REGION Network 3: I75.2 - Tank Vent Valve 1 Feedback Open (CV-441-A)
   // True = OPEN, False = NOT
   RUNG wire#powerrail
      Contact( "APT Tank Vent Valve 1 Feedback - Opened" )
      Coil( "20_TANKS_IP_DATA".RIO_07.FIRST_TANK.TANK_VENT_A_OPEN )
   END_RUNG
   // the same network as SCL:
   "20_TANKS_IP_DATA".RIO_07.FIRST_TANK.TANK_VENT_A_OPEN := "APT Tank Vent Valve 1 Feedback - Opened";
END_REGION

REGION Network 4: I75.3 - Tank Vent Valve 1 Feedback Closed (CV-441-A)
   // True = CLOSED, False = NOT
   RUNG wire#powerrail
      Contact( "APT Tank Vent Valve 1 Feedback - Closed" )
      Coil( "20_TANKS_IP_DATA".RIO_07.FIRST_TANK.TANK_VENT_A_CLSD )
   END_RUNG
   // the same network as SCL:
   "20_TANKS_IP_DATA".RIO_07.FIRST_TANK.TANK_VENT_A_CLSD := "APT Tank Vent Valve 1 Feedback - Closed";
END_REGION

REGION Network 5: I75.4 - Tank Vent Valve 2 Feedback Open (CV-441-B)
   // True = OPEN, False = NOT
   RUNG wire#powerrail
      Contact( "APT Tank Vent Valve 2 Feedback - Opened" )
      Coil( "20_TANKS_IP_DATA".RIO_07.FIRST_TANK.TANK_VENT_B_OPEN )
   END_RUNG
   // the same network as SCL:
   "20_TANKS_IP_DATA".RIO_07.FIRST_TANK.TANK_VENT_B_OPEN := "APT Tank Vent Valve 2 Feedback - Opened";
END_REGION

REGION Network 6: I75.5 - Tank Vent Valve 2 Feedback Closed (CV-441-B)
   // True = CLOSED, False = NOT
   RUNG wire#powerrail
      Contact( "APT Tank Vent Valve 2 Feedback - Closed" )
      Coil( "20_TANKS_IP_DATA".RIO_07.FIRST_TANK.TANK_VENT_B_CLSD )
   END_RUNG
   // the same network as SCL:
   "20_TANKS_IP_DATA".RIO_07.FIRST_TANK.TANK_VENT_B_CLSD := "APT Tank Vent Valve 2 Feedback - Closed";
END_REGION

REGION Network 7: I75.6 - Spare Input Destination Accesed from Warning FC
   // True = N/A, False = N/A
END_REGION

REGION Network 8: I75.7 - Spare Input
   // True = N/A, False = N/A
   RUNG wire#powerrail
      Contact( "RIO7_SPR_DI_175_7" )
      Coil( "20_TANKS_IP_DATA".RIO_07.FIRST_TANK.SPARE_DI_7 )
   END_RUNG
   // the same network as SCL:
   "20_TANKS_IP_DATA".RIO_07.FIRST_TANK.SPARE_DI_7 := "RIO7_SPR_DI_175_7";
END_REGION

REGION Network 9: I78.0 - Tank Level HIHI - (LS-425) - First Tank
   // True = OK, False = HIHI
   RUNG wire#powerrail
      I_Contact( "APT BWT Level High High Switch" )
      Coil( "20_TANKS_IP_DATA".RIO_07.FIRST_TANK.BWT_LEVEL_HIHI )
   END_RUNG
   // the same network as SCL:
   "20_TANKS_IP_DATA".RIO_07.FIRST_TANK.BWT_LEVEL_HIHI := NOT "APT BWT Level High High Switch";
END_REGION

REGION Network 10: I78.1 - Tank Group Pressure HIHI (PS-436)
   // True = OK, False = HIHI
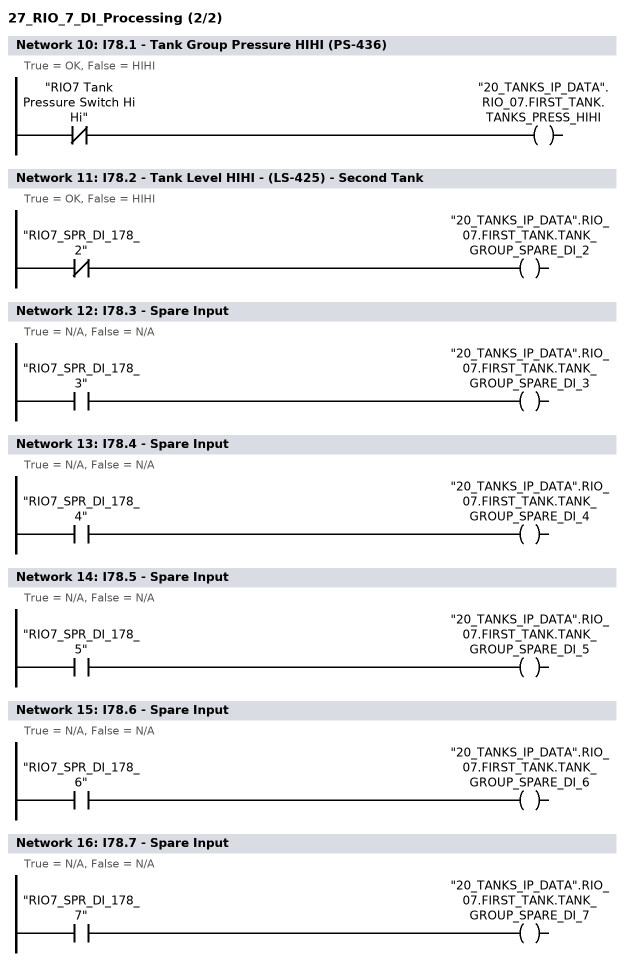
   RUNG wire#powerrail
      I_Contact( "RIO7 Tank Pressure Switch Hi Hi" )
      Coil( "20_TANKS_IP_DATA".RIO_07.FIRST_TANK.TANKS_PRESS_HIHI )
   END_RUNG
   // the same network as SCL:
   "20_TANKS_IP_DATA".RIO_07.FIRST_TANK.TANKS_PRESS_HIHI := NOT "RIO7 Tank Pressure Switch Hi Hi";
END_REGION

REGION Network 11: I78.2 - Tank Level HIHI - (LS-425) - Second Tank
   // True = OK, False = HIHI
   RUNG wire#powerrail
      I_Contact( "RIO7_SPR_DI_178_2" )
      Coil( "20_TANKS_IP_DATA".RIO_07.FIRST_TANK.TANK_GROUP_SPARE_DI_2 )
   END_RUNG
   // the same network as SCL:
   "20_TANKS_IP_DATA".RIO_07.FIRST_TANK.TANK_GROUP_SPARE_DI_2 := NOT "RIO7_SPR_DI_178_2";
END_REGION

REGION Network 12: I78.3 - Spare Input
   // True = N/A, False = N/A
   RUNG wire#powerrail
      Contact( "RIO7_SPR_DI_178_3" )
      Coil( "20_TANKS_IP_DATA".RIO_07.FIRST_TANK.TANK_GROUP_SPARE_DI_3 )
   END_RUNG
   // the same network as SCL:
   "20_TANKS_IP_DATA".RIO_07.FIRST_TANK.TANK_GROUP_SPARE_DI_3 := "RIO7_SPR_DI_178_3";
END_REGION

REGION Network 13: I78.4 - Spare Input
   // True = N/A, False = N/A
   RUNG wire#powerrail
      Contact( "RIO7_SPR_DI_178_4" )
      Coil( "20_TANKS_IP_DATA".RIO_07.FIRST_TANK.TANK_GROUP_SPARE_DI_4 )
   END_RUNG
   // the same network as SCL:
   "20_TANKS_IP_DATA".RIO_07.FIRST_TANK.TANK_GROUP_SPARE_DI_4 := "RIO7_SPR_DI_178_4";
END_REGION

REGION Network 14: I78.5 - Spare Input
   // True = N/A, False = N/A
   RUNG wire#powerrail
      Contact( "RIO7_SPR_DI_178_5" )
      Coil( "20_TANKS_IP_DATA".RIO_07.FIRST_TANK.TANK_GROUP_SPARE_DI_5 )
   END_RUNG
   // the same network as SCL:
   "20_TANKS_IP_DATA".RIO_07.FIRST_TANK.TANK_GROUP_SPARE_DI_5 := "RIO7_SPR_DI_178_5";
END_REGION

REGION Network 15: I78.6 - Spare Input
   // True = N/A, False = N/A
   RUNG wire#powerrail
      Contact( "RIO7_SPR_DI_178_6" )
      Coil( "20_TANKS_IP_DATA".RIO_07.FIRST_TANK.TANK_GROUP_SPARE_DI_6 )
   END_RUNG
   // the same network as SCL:
   "20_TANKS_IP_DATA".RIO_07.FIRST_TANK.TANK_GROUP_SPARE_DI_6 := "RIO7_SPR_DI_178_6";
END_REGION

REGION Network 16: I78.7 - Spare Input
   // True = N/A, False = N/A
   RUNG wire#powerrail
      Contact( "RIO7_SPR_DI_178_7" )
      Coil( "20_TANKS_IP_DATA".RIO_07.FIRST_TANK.TANK_GROUP_SPARE_DI_7 )
   END_RUNG
   // the same network as SCL:
   "20_TANKS_IP_DATA".RIO_07.FIRST_TANK.TANK_GROUP_SPARE_DI_7 := "RIO7_SPR_DI_178_7";
END_REGION
END_FUNCTION

FUNCTION "WBTs" : Void   // FC28, SCL
{ S7_Optimized_Access := 'TRUE' }
VERSION : 0.1
BEGIN
   "Data_From_WBT"."Level_FPT" := (INT_TO_REAL("IN_Level_FPT") / 1000.0) / "Data_From_WBT".Level_Max_FPT * 100.0;
   "Data_From_WBT"."Level_FPT m" := (INT_TO_REAL("IN_Level_FPT") / 1000.0);

   "Data_From_WBT"."Level_WBT_1S" := (INT_TO_REAL("IN_Level_WBT_1S") / 1000.0) /"Data_From_WBT".Level_Max_WBT_1S * 100.0;
   "Data_From_WBT"."Level_WBT_1P" := (INT_TO_REAL("IN_Level_WBT_1P") / 1000.0) / "Data_From_WBT".Level_Max_WBT_1P * 100.0;
   "Data_From_WBT"."Level_WBT_1S m" := (INT_TO_REAL("IN_Level_WBT_1S") / 1000.0);
   "Data_From_WBT"."Level_WBT_1P m" := (INT_TO_REAL("IN_Level_WBT_1P") / 1000.0);

   "Data_From_WBT"."Level_WBT_2S" := (INT_TO_REAL("IN_Level_WBT_2S") / 1000.0) / "Data_From_WBT".Level_Max_WBT_2S * 100.0;
   "Data_From_WBT"."Level_WBT_2P" := (INT_TO_REAL("IN_Level_WBT_2P") / 1000.0) / "Data_From_WBT".Level_Max_WBT_2P * 100.0;
   "Data_From_WBT"."Level_WBT_2S m":= (INT_TO_REAL("IN_Level_WBT_2S") / 1000.0);
   "Data_From_WBT"."Level_WBT_2P m" := (INT_TO_REAL("IN_Level_WBT_2P") / 1000.0);

   "Data_From_WBT"."Level_WBT_3S" := (INT_TO_REAL("IN_Level_WBT_3S") / 1000.0) / "Data_From_WBT".Level_Max_WBT_3S * 100.0;
   "Data_From_WBT"."Level_WBT_3P" := (INT_TO_REAL("IN_Level_WBT_3P") / 1000.0) / "Data_From_WBT".Level_Max_WBT_3P * 100.0;
   "Data_From_WBT"."Level_WBT_3S m" := (INT_TO_REAL("IN_Level_WBT_3S") / 1000.0);
   "Data_From_WBT"."Level_WBT_3P m" := (INT_TO_REAL("IN_Level_WBT_3P") / 1000.0);

   "Data_From_WBT"."Level_WBT_4S" := (INT_TO_REAL("IN_Level_WBT_4S") / 1000.0) / "Data_From_WBT".Level_Max_WBT_4S * 100.0;
   "Data_From_WBT"."Level_WBT_4P" := (INT_TO_REAL("IN_Level_WBT_4P") / 1000.0) / "Data_From_WBT".Level_Max_WBT_4P * 100.0;
   "Data_From_WBT"."Level_WBT_4S m" := (INT_TO_REAL("IN_Level_WBT_4S") / 1000.0);
   "Data_From_WBT"."Level_WBT_4P m" := (INT_TO_REAL("IN_Level_WBT_4P") / 1000.0);

   "Data_From_WBT"."Level_WBT_5S" := (INT_TO_REAL("IN_Level_WBT_5S") / 1000.0) / "Data_From_WBT".Level_Max_WBT_5S * 100.0;
   "Data_From_WBT"."Level_WBT_5P" := (INT_TO_REAL("IN_Level_WBT_5P") / 1000.0) / "Data_From_WBT".Level_Max_WBT_5P * 100.0;
   "Data_From_WBT"."Level_WBT_5S m" := (INT_TO_REAL("IN_Level_WBT_5S") / 1000.0);
   "Data_From_WBT"."Level_WBT_5P m" := (INT_TO_REAL("IN_Level_WBT_5P") / 1000.0);

   "Data_From_WBT"."Level_WBT_6S" := (INT_TO_REAL("IN_Level_WBT_6S") / 1000.0) / "Data_From_WBT".Level_Max_WBT_6S * 100.0;
   "Data_From_WBT"."Level_WBT_6P" := (INT_TO_REAL("IN_Level_WBT_6P") / 1000.0) / "Data_From_WBT".Level_Max_WBT_6P * 100.0;
   "Data_From_WBT"."Level_WBT_6S m" := (INT_TO_REAL("IN_Level_WBT_6S") / 1000.0);
   "Data_From_WBT"."Level_WBT_6P m" := (INT_TO_REAL("IN_Level_WBT_6P") / 1000.0);

   "Data_From_WBT"."Level_APT" := (INT_TO_REAL("IN_Level_APT") / 1000.0) / "Data_From_WBT".Level_Max_APT * 100.0;
   "Data_From_WBT"."Level_APT m" := (INT_TO_REAL("IN_Level_APT") / 1000.0);
END_FUNCTION

FUNCTION "31_RIO_1_AI_Processing" : Void   // FC31, LAD
TITLE = Analogue Input Processing (Tank 1 = FPT, Tank 2 = 1P, Tank 3 = 1S)
{ S7_Optimized_Access := 'TRUE' }
AUTHOR : JRS
VERSION : 0.1
// To process raw inputs prior to code use
BEGIN

REGION Network 1: IW100 - USD Flow (FIT-418) - Tank #1
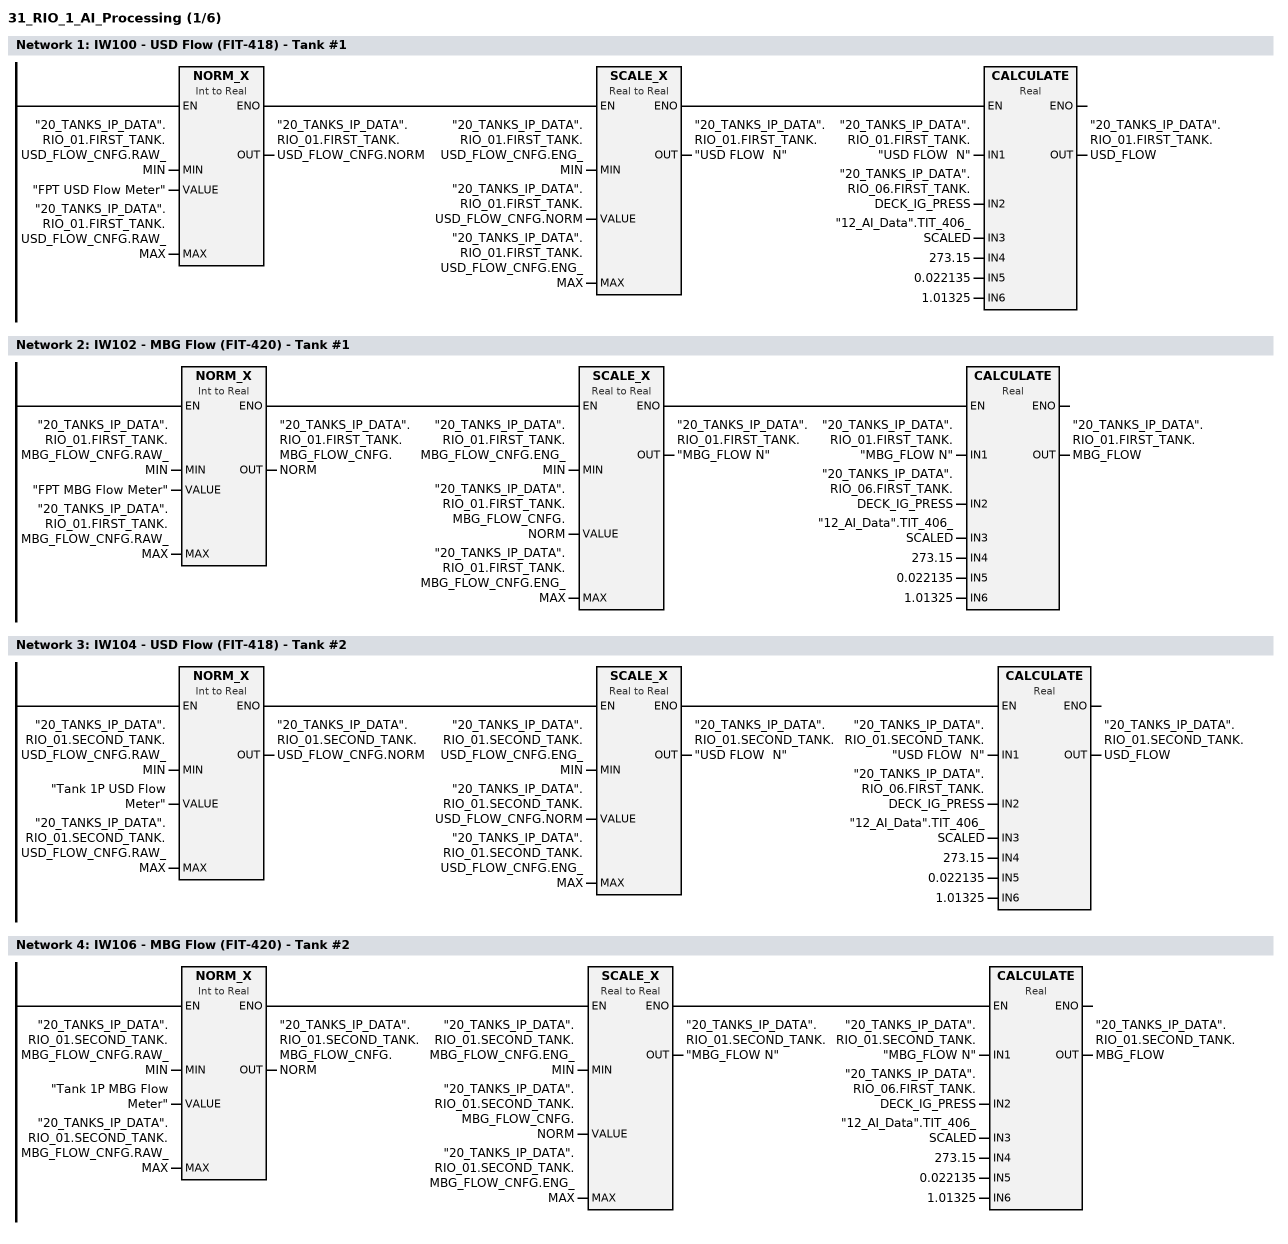
   RUNG wire#powerrail
      { S7_Templates := "[SrcType := Int, DestType := Real]" } Normalize(min := "20_TANKS_IP_DATA".RIO_01.FIRST_TANK.USD_FLOW_CNFG.RAW_MIN, value := "FPT USD Flow Meter", max := "20_TANKS_IP_DATA".RIO_01.FIRST_TANK.USD_FLOW_CNFG.RAW_MAX, out => "20_TANKS_IP_DATA".RIO_01.FIRST_TANK.USD_FLOW_CNFG.NORM)
      { S7_Templates := "[SrcType := Real, DestType := Real]" } Scale(min := "20_TANKS_IP_DATA".RIO_01.FIRST_TANK.USD_FLOW_CNFG.ENG_MIN, value := "20_TANKS_IP_DATA".RIO_01.FIRST_TANK.USD_FLOW_CNFG.NORM, max := "20_TANKS_IP_DATA".RIO_01.FIRST_TANK.USD_FLOW_CNFG.ENG_MAX, out => "20_TANKS_IP_DATA".RIO_01.FIRST_TANK."USD FLOW  N")
      { S7_Templates := "SrcType := Real"; S7_Expression := "IN1*(IN2+IN6)/IN6*IN4/(IN3+IN4)" } Calculate(in1 := "20_TANKS_IP_DATA".RIO_01.FIRST_TANK."USD FLOW  N", in2 := "20_TANKS_IP_DATA".RIO_06.FIRST_TANK.DECK_IG_PRESS, in3 := "12_AI_Data".TIT_406_SCALED, in4 := 273.15, in5 := 0.022135, in6 := 1.01325, out => "20_TANKS_IP_DATA".RIO_01.FIRST_TANK.USD_FLOW)
   END_RUNG
   // the same network as SCL:
   "20_TANKS_IP_DATA".RIO_01.FIRST_TANK.USD_FLOW_CNFG.NORM := NORM_X(MIN := "20_TANKS_IP_DATA".RIO_01.FIRST_TANK.USD_FLOW_CNFG.RAW_MIN, VALUE := "FPT USD Flow Meter", MAX := "20_TANKS_IP_DATA".RIO_01.FIRST_TANK.USD_FLOW_CNFG.RAW_MAX);
   "20_TANKS_IP_DATA".RIO_01.FIRST_TANK."USD FLOW  N" := SCALE_X(MIN := "20_TANKS_IP_DATA".RIO_01.FIRST_TANK.USD_FLOW_CNFG.ENG_MIN, VALUE := "20_TANKS_IP_DATA".RIO_01.FIRST_TANK.USD_FLOW_CNFG.NORM, MAX := "20_TANKS_IP_DATA".RIO_01.FIRST_TANK.USD_FLOW_CNFG.ENG_MAX);
   "20_TANKS_IP_DATA".RIO_01.FIRST_TANK.USD_FLOW := "20_TANKS_IP_DATA".RIO_01.FIRST_TANK."USD FLOW  N"*("20_TANKS_IP_DATA".RIO_06.FIRST_TANK.DECK_IG_PRESS+1.01325)/1.01325*273.15/("12_AI_Data".TIT_406_SCALED+273.15);
END_REGION

REGION Network 2: IW102 - MBG Flow (FIT-420) - Tank #1
   RUNG wire#powerrail
      { S7_Templates := "[SrcType := Int, DestType := Real]" } Normalize(min := "20_TANKS_IP_DATA".RIO_01.FIRST_TANK.MBG_FLOW_CNFG.RAW_MIN, value := "FPT MBG Flow Meter", max := "20_TANKS_IP_DATA".RIO_01.FIRST_TANK.MBG_FLOW_CNFG.RAW_MAX, out => "20_TANKS_IP_DATA".RIO_01.FIRST_TANK.MBG_FLOW_CNFG.NORM)
      { S7_Templates := "[SrcType := Real, DestType := Real]" } Scale(min := "20_TANKS_IP_DATA".RIO_01.FIRST_TANK.MBG_FLOW_CNFG.ENG_MIN, value := "20_TANKS_IP_DATA".RIO_01.FIRST_TANK.MBG_FLOW_CNFG.NORM, max := "20_TANKS_IP_DATA".RIO_01.FIRST_TANK.MBG_FLOW_CNFG.ENG_MAX, out => "20_TANKS_IP_DATA".RIO_01.FIRST_TANK."MBG_FLOW N")
      { S7_Templates := "SrcType := Real"; S7_Expression := "IN1*(IN2+IN6)/IN6*IN4/(IN3+IN4)" } Calculate(in1 := "20_TANKS_IP_DATA".RIO_01.FIRST_TANK."MBG_FLOW N", in2 := "20_TANKS_IP_DATA".RIO_06.FIRST_TANK.DECK_IG_PRESS, in3 := "12_AI_Data".TIT_406_SCALED, in4 := 273.15, in5 := 0.022135, in6 := 1.01325, out => "20_TANKS_IP_DATA".RIO_01.FIRST_TANK.MBG_FLOW)
   END_RUNG
   // the same network as SCL:
   "20_TANKS_IP_DATA".RIO_01.FIRST_TANK.MBG_FLOW_CNFG.NORM := NORM_X(MIN := "20_TANKS_IP_DATA".RIO_01.FIRST_TANK.MBG_FLOW_CNFG.RAW_MIN, VALUE := "FPT MBG Flow Meter", MAX := "20_TANKS_IP_DATA".RIO_01.FIRST_TANK.MBG_FLOW_CNFG.RAW_MAX);
   "20_TANKS_IP_DATA".RIO_01.FIRST_TANK."MBG_FLOW N" := SCALE_X(MIN := "20_TANKS_IP_DATA".RIO_01.FIRST_TANK.MBG_FLOW_CNFG.ENG_MIN, VALUE := "20_TANKS_IP_DATA".RIO_01.FIRST_TANK.MBG_FLOW_CNFG.NORM, MAX := "20_TANKS_IP_DATA".RIO_01.FIRST_TANK.MBG_FLOW_CNFG.ENG_MAX);
   "20_TANKS_IP_DATA".RIO_01.FIRST_TANK.MBG_FLOW := "20_TANKS_IP_DATA".RIO_01.FIRST_TANK."MBG_FLOW N"*("20_TANKS_IP_DATA".RIO_06.FIRST_TANK.DECK_IG_PRESS+1.01325)/1.01325*273.15/("12_AI_Data".TIT_406_SCALED+273.15);
END_REGION

REGION Network 3: IW104 - USD Flow (FIT-418) - Tank #2
   RUNG wire#powerrail
      { S7_Templates := "[SrcType := Int, DestType := Real]" } Normalize(min := "20_TANKS_IP_DATA".RIO_01.SECOND_TANK.USD_FLOW_CNFG.RAW_MIN, value := "Tank 1P USD Flow Meter", max := "20_TANKS_IP_DATA".RIO_01.SECOND_TANK.USD_FLOW_CNFG.RAW_MAX, out => "20_TANKS_IP_DATA".RIO_01.SECOND_TANK.USD_FLOW_CNFG.NORM)
      { S7_Templates := "[SrcType := Real, DestType := Real]" } Scale(min := "20_TANKS_IP_DATA".RIO_01.SECOND_TANK.USD_FLOW_CNFG.ENG_MIN, value := "20_TANKS_IP_DATA".RIO_01.SECOND_TANK.USD_FLOW_CNFG.NORM, max := "20_TANKS_IP_DATA".RIO_01.SECOND_TANK.USD_FLOW_CNFG.ENG_MAX, out => "20_TANKS_IP_DATA".RIO_01.SECOND_TANK."USD FLOW  N")
      { S7_Templates := "SrcType := Real"; S7_Expression := "IN1*(IN2+IN6)/IN6*IN4/(IN3+IN4)" } Calculate(in1 := "20_TANKS_IP_DATA".RIO_01.SECOND_TANK."USD FLOW  N", in2 := "20_TANKS_IP_DATA".RIO_06.FIRST_TANK.DECK_IG_PRESS, in3 := "12_AI_Data".TIT_406_SCALED, in4 := 273.15, in5 := 0.022135, in6 := 1.01325, out => "20_TANKS_IP_DATA".RIO_01.SECOND_TANK.USD_FLOW)
   END_RUNG
   // the same network as SCL:
   "20_TANKS_IP_DATA".RIO_01.SECOND_TANK.USD_FLOW_CNFG.NORM := NORM_X(MIN := "20_TANKS_IP_DATA".RIO_01.SECOND_TANK.USD_FLOW_CNFG.RAW_MIN, VALUE := "Tank 1P USD Flow Meter", MAX := "20_TANKS_IP_DATA".RIO_01.SECOND_TANK.USD_FLOW_CNFG.RAW_MAX);
   "20_TANKS_IP_DATA".RIO_01.SECOND_TANK."USD FLOW  N" := SCALE_X(MIN := "20_TANKS_IP_DATA".RIO_01.SECOND_TANK.USD_FLOW_CNFG.ENG_MIN, VALUE := "20_TANKS_IP_DATA".RIO_01.SECOND_TANK.USD_FLOW_CNFG.NORM, MAX := "20_TANKS_IP_DATA".RIO_01.SECOND_TANK.USD_FLOW_CNFG.ENG_MAX);
   "20_TANKS_IP_DATA".RIO_01.SECOND_TANK.USD_FLOW := "20_TANKS_IP_DATA".RIO_01.SECOND_TANK."USD FLOW  N"*("20_TANKS_IP_DATA".RIO_06.FIRST_TANK.DECK_IG_PRESS+1.01325)/1.01325*273.15/("12_AI_Data".TIT_406_SCALED+273.15);
END_REGION

REGION Network 4: IW106 - MBG Flow (FIT-420) - Tank #2
   RUNG wire#powerrail
      { S7_Templates := "[SrcType := Int, DestType := Real]" } Normalize(min := "20_TANKS_IP_DATA".RIO_01.SECOND_TANK.MBG_FLOW_CNFG.RAW_MIN, value := "Tank 1P MBG Flow Meter", max := "20_TANKS_IP_DATA".RIO_01.SECOND_TANK.MBG_FLOW_CNFG.RAW_MAX, out => "20_TANKS_IP_DATA".RIO_01.SECOND_TANK.MBG_FLOW_CNFG.NORM)
      { S7_Templates := "[SrcType := Real, DestType := Real]" } Scale(min := "20_TANKS_IP_DATA".RIO_01.SECOND_TANK.MBG_FLOW_CNFG.ENG_MIN, value := "20_TANKS_IP_DATA".RIO_01.SECOND_TANK.MBG_FLOW_CNFG.NORM, max := "20_TANKS_IP_DATA".RIO_01.SECOND_TANK.MBG_FLOW_CNFG.ENG_MAX, out => "20_TANKS_IP_DATA".RIO_01.SECOND_TANK."MBG_FLOW N")
      { S7_Templates := "SrcType := Real"; S7_Expression := "IN1*(IN2+IN6)/IN6*IN4/(IN3+IN4)" } Calculate(in1 := "20_TANKS_IP_DATA".RIO_01.SECOND_TANK."MBG_FLOW N", in2 := "20_TANKS_IP_DATA".RIO_06.FIRST_TANK.DECK_IG_PRESS, in3 := "12_AI_Data".TIT_406_SCALED, in4 := 273.15, in5 := 0.022135, in6 := 1.01325, out => "20_TANKS_IP_DATA".RIO_01.SECOND_TANK.MBG_FLOW)
   END_RUNG
   // the same network as SCL:
   "20_TANKS_IP_DATA".RIO_01.SECOND_TANK.MBG_FLOW_CNFG.NORM := NORM_X(MIN := "20_TANKS_IP_DATA".RIO_01.SECOND_TANK.MBG_FLOW_CNFG.RAW_MIN, VALUE := "Tank 1P MBG Flow Meter", MAX := "20_TANKS_IP_DATA".RIO_01.SECOND_TANK.MBG_FLOW_CNFG.RAW_MAX);
   "20_TANKS_IP_DATA".RIO_01.SECOND_TANK."MBG_FLOW N" := SCALE_X(MIN := "20_TANKS_IP_DATA".RIO_01.SECOND_TANK.MBG_FLOW_CNFG.ENG_MIN, VALUE := "20_TANKS_IP_DATA".RIO_01.SECOND_TANK.MBG_FLOW_CNFG.NORM, MAX := "20_TANKS_IP_DATA".RIO_01.SECOND_TANK.MBG_FLOW_CNFG.ENG_MAX);
   "20_TANKS_IP_DATA".RIO_01.SECOND_TANK.MBG_FLOW := "20_TANKS_IP_DATA".RIO_01.SECOND_TANK."MBG_FLOW N"*("20_TANKS_IP_DATA".RIO_06.FIRST_TANK.DECK_IG_PRESS+1.01325)/1.01325*273.15/("12_AI_Data".TIT_406_SCALED+273.15);
END_REGION

REGION Network 5: IW108 - USD Flow (FIT-418) - Tank #3
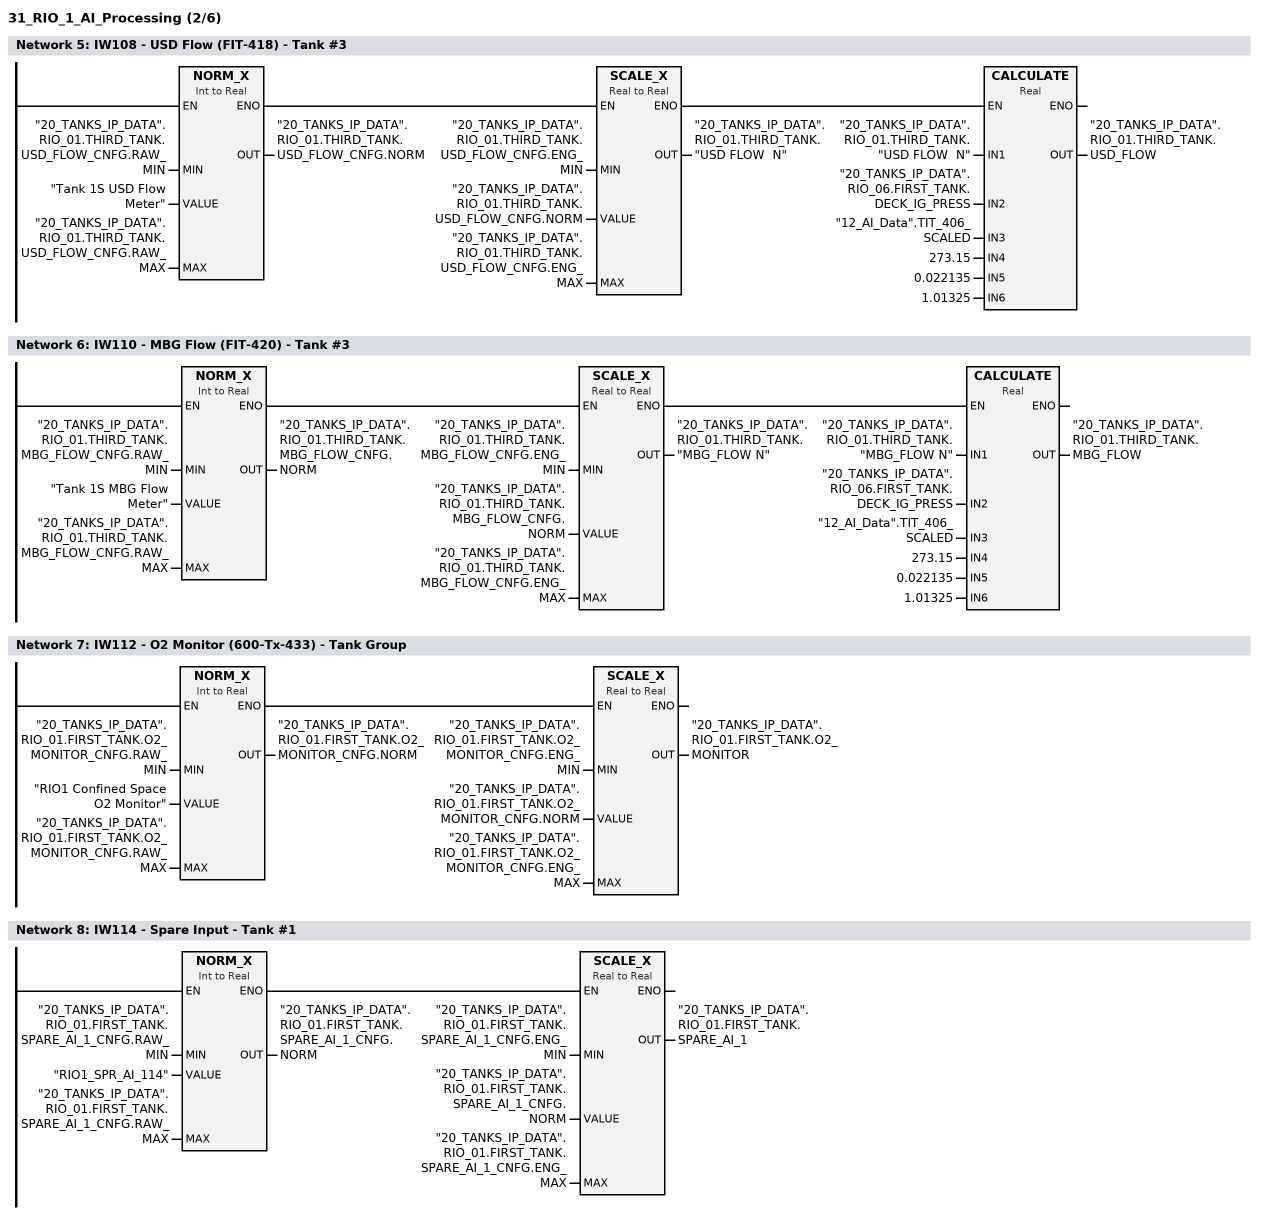
   RUNG wire#powerrail
      { S7_Templates := "[SrcType := Int, DestType := Real]" } Normalize(min := "20_TANKS_IP_DATA".RIO_01.THIRD_TANK.USD_FLOW_CNFG.RAW_MIN, value := "Tank 1S USD Flow Meter", max := "20_TANKS_IP_DATA".RIO_01.THIRD_TANK.USD_FLOW_CNFG.RAW_MAX, out => "20_TANKS_IP_DATA".RIO_01.THIRD_TANK.USD_FLOW_CNFG.NORM)
      { S7_Templates := "[SrcType := Real, DestType := Real]" } Scale(min := "20_TANKS_IP_DATA".RIO_01.THIRD_TANK.USD_FLOW_CNFG.ENG_MIN, value := "20_TANKS_IP_DATA".RIO_01.THIRD_TANK.USD_FLOW_CNFG.NORM, max := "20_TANKS_IP_DATA".RIO_01.THIRD_TANK.USD_FLOW_CNFG.ENG_MAX, out => "20_TANKS_IP_DATA".RIO_01.THIRD_TANK."USD FLOW  N")
      { S7_Templates := "SrcType := Real"; S7_Expression := "IN1*(IN2+IN6)/IN6*IN4/(IN3+IN4)" } Calculate(in1 := "20_TANKS_IP_DATA".RIO_01.THIRD_TANK."USD FLOW  N", in2 := "20_TANKS_IP_DATA".RIO_06.FIRST_TANK.DECK_IG_PRESS, in3 := "12_AI_Data".TIT_406_SCALED, in4 := 273.15, in5 := 0.022135, in6 := 1.01325, out => "20_TANKS_IP_DATA".RIO_01.THIRD_TANK.USD_FLOW)
   END_RUNG
   // the same network as SCL:
   "20_TANKS_IP_DATA".RIO_01.THIRD_TANK.USD_FLOW_CNFG.NORM := NORM_X(MIN := "20_TANKS_IP_DATA".RIO_01.THIRD_TANK.USD_FLOW_CNFG.RAW_MIN, VALUE := "Tank 1S USD Flow Meter", MAX := "20_TANKS_IP_DATA".RIO_01.THIRD_TANK.USD_FLOW_CNFG.RAW_MAX);
   "20_TANKS_IP_DATA".RIO_01.THIRD_TANK."USD FLOW  N" := SCALE_X(MIN := "20_TANKS_IP_DATA".RIO_01.THIRD_TANK.USD_FLOW_CNFG.ENG_MIN, VALUE := "20_TANKS_IP_DATA".RIO_01.THIRD_TANK.USD_FLOW_CNFG.NORM, MAX := "20_TANKS_IP_DATA".RIO_01.THIRD_TANK.USD_FLOW_CNFG.ENG_MAX);
   "20_TANKS_IP_DATA".RIO_01.THIRD_TANK.USD_FLOW := "20_TANKS_IP_DATA".RIO_01.THIRD_TANK."USD FLOW  N"*("20_TANKS_IP_DATA".RIO_06.FIRST_TANK.DECK_IG_PRESS+1.01325)/1.01325*273.15/("12_AI_Data".TIT_406_SCALED+273.15);
END_REGION

REGION Network 6: IW110 - MBG Flow (FIT-420) - Tank #3
   RUNG wire#powerrail
      { S7_Templates := "[SrcType := Int, DestType := Real]" } Normalize(min := "20_TANKS_IP_DATA".RIO_01.THIRD_TANK.MBG_FLOW_CNFG.RAW_MIN, value := "Tank 1S MBG Flow Meter", max := "20_TANKS_IP_DATA".RIO_01.THIRD_TANK.MBG_FLOW_CNFG.RAW_MAX, out => "20_TANKS_IP_DATA".RIO_01.THIRD_TANK.MBG_FLOW_CNFG.NORM)
      { S7_Templates := "[SrcType := Real, DestType := Real]" } Scale(min := "20_TANKS_IP_DATA".RIO_01.THIRD_TANK.MBG_FLOW_CNFG.ENG_MIN, value := "20_TANKS_IP_DATA".RIO_01.THIRD_TANK.MBG_FLOW_CNFG.NORM, max := "20_TANKS_IP_DATA".RIO_01.THIRD_TANK.MBG_FLOW_CNFG.ENG_MAX, out => "20_TANKS_IP_DATA".RIO_01.THIRD_TANK."MBG_FLOW N")
      { S7_Templates := "SrcType := Real"; S7_Expression := "IN1*(IN2+IN6)/IN6*IN4/(IN3+IN4)" } Calculate(in1 := "20_TANKS_IP_DATA".RIO_01.THIRD_TANK."MBG_FLOW N", in2 := "20_TANKS_IP_DATA".RIO_06.FIRST_TANK.DECK_IG_PRESS, in3 := "12_AI_Data".TIT_406_SCALED, in4 := 273.15, in5 := 0.022135, in6 := 1.01325, out => "20_TANKS_IP_DATA".RIO_01.THIRD_TANK.MBG_FLOW)
   END_RUNG
   // the same network as SCL:
   "20_TANKS_IP_DATA".RIO_01.THIRD_TANK.MBG_FLOW_CNFG.NORM := NORM_X(MIN := "20_TANKS_IP_DATA".RIO_01.THIRD_TANK.MBG_FLOW_CNFG.RAW_MIN, VALUE := "Tank 1S MBG Flow Meter", MAX := "20_TANKS_IP_DATA".RIO_01.THIRD_TANK.MBG_FLOW_CNFG.RAW_MAX);
   "20_TANKS_IP_DATA".RIO_01.THIRD_TANK."MBG_FLOW N" := SCALE_X(MIN := "20_TANKS_IP_DATA".RIO_01.THIRD_TANK.MBG_FLOW_CNFG.ENG_MIN, VALUE := "20_TANKS_IP_DATA".RIO_01.THIRD_TANK.MBG_FLOW_CNFG.NORM, MAX := "20_TANKS_IP_DATA".RIO_01.THIRD_TANK.MBG_FLOW_CNFG.ENG_MAX);
   "20_TANKS_IP_DATA".RIO_01.THIRD_TANK.MBG_FLOW := "20_TANKS_IP_DATA".RIO_01.THIRD_TANK."MBG_FLOW N"*("20_TANKS_IP_DATA".RIO_06.FIRST_TANK.DECK_IG_PRESS+1.01325)/1.01325*273.15/("12_AI_Data".TIT_406_SCALED+273.15);
END_REGION

REGION Network 7: IW112 - O2 Monitor (600-Tx-433) - Tank Group
   RUNG wire#powerrail
      { S7_Templates := "[SrcType := Int, DestType := Real]" } Normalize(min := "20_TANKS_IP_DATA".RIO_01.FIRST_TANK.O2_MONITOR_CNFG.RAW_MIN, value := "RIO1 Confined Space O2 Monitor", max := "20_TANKS_IP_DATA".RIO_01.FIRST_TANK.O2_MONITOR_CNFG.RAW_MAX, out => "20_TANKS_IP_DATA".RIO_01.FIRST_TANK.O2_MONITOR_CNFG.NORM)
      { S7_Templates := "[SrcType := Real, DestType := Real]" } Scale(min := "20_TANKS_IP_DATA".RIO_01.FIRST_TANK.O2_MONITOR_CNFG.ENG_MIN, value := "20_TANKS_IP_DATA".RIO_01.FIRST_TANK.O2_MONITOR_CNFG.NORM, max := "20_TANKS_IP_DATA".RIO_01.FIRST_TANK.O2_MONITOR_CNFG.ENG_MAX, out => "20_TANKS_IP_DATA".RIO_01.FIRST_TANK.O2_MONITOR)
   END_RUNG
   // the same network as SCL:
   "20_TANKS_IP_DATA".RIO_01.FIRST_TANK.O2_MONITOR_CNFG.NORM := NORM_X(MIN := "20_TANKS_IP_DATA".RIO_01.FIRST_TANK.O2_MONITOR_CNFG.RAW_MIN, VALUE := "RIO1 Confined Space O2 Monitor", MAX := "20_TANKS_IP_DATA".RIO_01.FIRST_TANK.O2_MONITOR_CNFG.RAW_MAX);
   "20_TANKS_IP_DATA".RIO_01.FIRST_TANK.O2_MONITOR := SCALE_X(MIN := "20_TANKS_IP_DATA".RIO_01.FIRST_TANK.O2_MONITOR_CNFG.ENG_MIN, VALUE := "20_TANKS_IP_DATA".RIO_01.FIRST_TANK.O2_MONITOR_CNFG.NORM, MAX := "20_TANKS_IP_DATA".RIO_01.FIRST_TANK.O2_MONITOR_CNFG.ENG_MAX);
END_REGION

REGION Network 8: IW114 - Spare Input - Tank #1
   RUNG wire#powerrail
      { S7_Templates := "[SrcType := Int, DestType := Real]" } Normalize(min := "20_TANKS_IP_DATA".RIO_01.FIRST_TANK.SPARE_AI_1_CNFG.RAW_MIN, value := "RIO1_SPR_AI_114", max := "20_TANKS_IP_DATA".RIO_01.FIRST_TANK.SPARE_AI_1_CNFG.RAW_MAX, out => "20_TANKS_IP_DATA".RIO_01.FIRST_TANK.SPARE_AI_1_CNFG.NORM)
      { S7_Templates := "[SrcType := Real, DestType := Real]" } Scale(min := "20_TANKS_IP_DATA".RIO_01.FIRST_TANK.SPARE_AI_1_CNFG.ENG_MIN, value := "20_TANKS_IP_DATA".RIO_01.FIRST_TANK.SPARE_AI_1_CNFG.NORM, max := "20_TANKS_IP_DATA".RIO_01.FIRST_TANK.SPARE_AI_1_CNFG.ENG_MAX, out => "20_TANKS_IP_DATA".RIO_01.FIRST_TANK.SPARE_AI_1)
   END_RUNG
   // the same network as SCL:
   "20_TANKS_IP_DATA".RIO_01.FIRST_TANK.SPARE_AI_1_CNFG.NORM := NORM_X(MIN := "20_TANKS_IP_DATA".RIO_01.FIRST_TANK.SPARE_AI_1_CNFG.RAW_MIN, VALUE := "RIO1_SPR_AI_114", MAX := "20_TANKS_IP_DATA".RIO_01.FIRST_TANK.SPARE_AI_1_CNFG.RAW_MAX);
   "20_TANKS_IP_DATA".RIO_01.FIRST_TANK.SPARE_AI_1 := SCALE_X(MIN := "20_TANKS_IP_DATA".RIO_01.FIRST_TANK.SPARE_AI_1_CNFG.ENG_MIN, VALUE := "20_TANKS_IP_DATA".RIO_01.FIRST_TANK.SPARE_AI_1_CNFG.NORM, MAX := "20_TANKS_IP_DATA".RIO_01.FIRST_TANK.SPARE_AI_1_CNFG.ENG_MAX);
END_REGION

REGION Network 9: IW116 - Deck Main IG Pressure (PT-415) - Tank Group
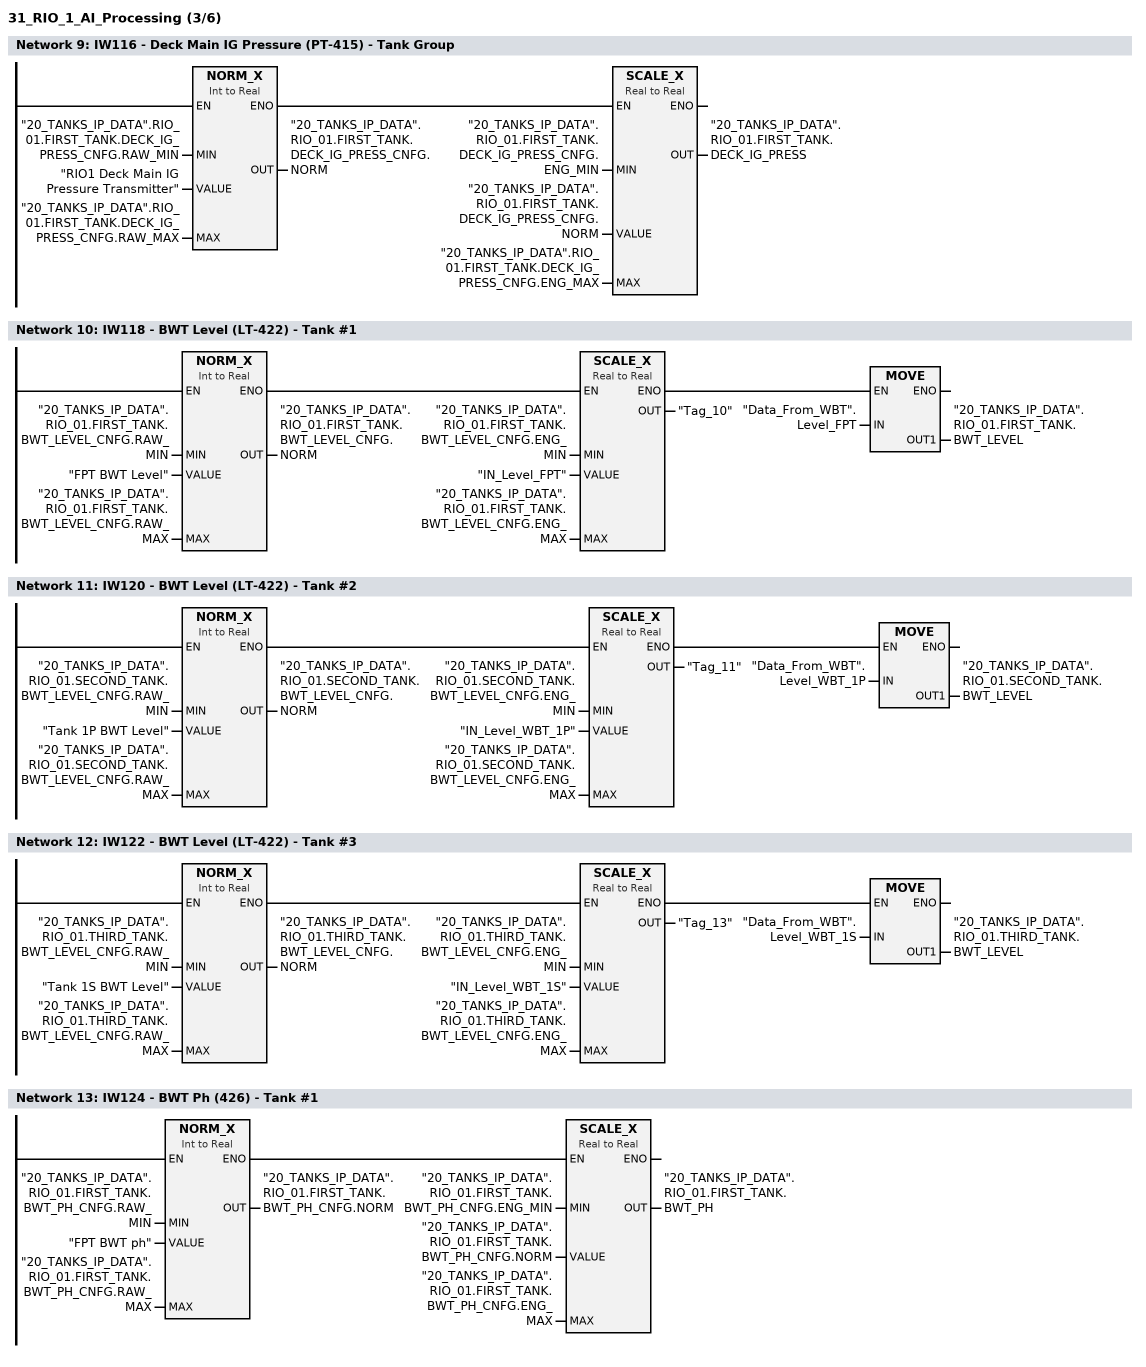
   RUNG wire#powerrail
      { S7_Templates := "[SrcType := Int, DestType := Real]" } Normalize(min := "20_TANKS_IP_DATA".RIO_01.FIRST_TANK.DECK_IG_PRESS_CNFG.RAW_MIN, value := "RIO1 Deck Main IG Pressure Transmitter", max := "20_TANKS_IP_DATA".RIO_01.FIRST_TANK.DECK_IG_PRESS_CNFG.RAW_MAX, out => "20_TANKS_IP_DATA".RIO_01.FIRST_TANK.DECK_IG_PRESS_CNFG.NORM)
      { S7_Templates := "[SrcType := Real, DestType := Real]" } Scale(min := "20_TANKS_IP_DATA".RIO_01.FIRST_TANK.DECK_IG_PRESS_CNFG.ENG_MIN, value := "20_TANKS_IP_DATA".RIO_01.FIRST_TANK.DECK_IG_PRESS_CNFG.NORM, max := "20_TANKS_IP_DATA".RIO_01.FIRST_TANK.DECK_IG_PRESS_CNFG.ENG_MAX, out => "20_TANKS_IP_DATA".RIO_01.FIRST_TANK.DECK_IG_PRESS)
   END_RUNG
   // the same network as SCL:
   "20_TANKS_IP_DATA".RIO_01.FIRST_TANK.DECK_IG_PRESS_CNFG.NORM := NORM_X(MIN := "20_TANKS_IP_DATA".RIO_01.FIRST_TANK.DECK_IG_PRESS_CNFG.RAW_MIN, VALUE := "RIO1 Deck Main IG Pressure Transmitter", MAX := "20_TANKS_IP_DATA".RIO_01.FIRST_TANK.DECK_IG_PRESS_CNFG.RAW_MAX);
   "20_TANKS_IP_DATA".RIO_01.FIRST_TANK.DECK_IG_PRESS := SCALE_X(MIN := "20_TANKS_IP_DATA".RIO_01.FIRST_TANK.DECK_IG_PRESS_CNFG.ENG_MIN, VALUE := "20_TANKS_IP_DATA".RIO_01.FIRST_TANK.DECK_IG_PRESS_CNFG.NORM, MAX := "20_TANKS_IP_DATA".RIO_01.FIRST_TANK.DECK_IG_PRESS_CNFG.ENG_MAX);
END_REGION

REGION Network 10: IW118 - BWT Level (LT-422) - Tank #1
   RUNG wire#powerrail
      { S7_Templates := "[SrcType := Int, DestType := Real]" } Normalize(min := "20_TANKS_IP_DATA".RIO_01.FIRST_TANK.BWT_LEVEL_CNFG.RAW_MIN, value := "FPT BWT Level", max := "20_TANKS_IP_DATA".RIO_01.FIRST_TANK.BWT_LEVEL_CNFG.RAW_MAX, out => "20_TANKS_IP_DATA".RIO_01.FIRST_TANK.BWT_LEVEL_CNFG.NORM)
      { S7_Templates := "[SrcType := Real, DestType := Real]" } Scale(min := "20_TANKS_IP_DATA".RIO_01.FIRST_TANK.BWT_LEVEL_CNFG.ENG_MIN, value := "IN_Level_FPT", max := "20_TANKS_IP_DATA".RIO_01.FIRST_TANK.BWT_LEVEL_CNFG.ENG_MAX, out => "Tag_10")
      Move(in := "Data_From_WBT".Level_FPT, out1 => "20_TANKS_IP_DATA".RIO_01.FIRST_TANK.BWT_LEVEL)
   END_RUNG
   // the same network as SCL:
   "20_TANKS_IP_DATA".RIO_01.FIRST_TANK.BWT_LEVEL_CNFG.NORM := NORM_X(MIN := "20_TANKS_IP_DATA".RIO_01.FIRST_TANK.BWT_LEVEL_CNFG.RAW_MIN, VALUE := "FPT BWT Level", MAX := "20_TANKS_IP_DATA".RIO_01.FIRST_TANK.BWT_LEVEL_CNFG.RAW_MAX);
   "Tag_10" := SCALE_X(MIN := "20_TANKS_IP_DATA".RIO_01.FIRST_TANK.BWT_LEVEL_CNFG.ENG_MIN, VALUE := "IN_Level_FPT", MAX := "20_TANKS_IP_DATA".RIO_01.FIRST_TANK.BWT_LEVEL_CNFG.ENG_MAX);
   "20_TANKS_IP_DATA".RIO_01.FIRST_TANK.BWT_LEVEL := "Data_From_WBT".Level_FPT;
END_REGION
